   hmiStns[3].wip[6].pnCode[4] := 0;
   hmiStns[3].wip[6].pnCode[5] := 0;
   hmiStns[3].wip[6].pnCode[6] := 197000;
   hmiStns[3].wip[6].pnCode[7] := 179000;
   hmiStns[3].wip[7].wipCode := -1;
   hmiStns[3].wip[7].pnCode[0] := 0;
   hmiStns[3].wip[7].pnCode[1] := 243000;
   hmiStns[3].wip[7].pnCode[2] := 0;
   hmiStns[3].wip[7].pnCode[3] := 199000;
   hmiStns[3].wip[7].pnCode[4] := 0;
   hmiStns[3].wip[7].pnCode[5] := 0;
   hmiStns[3].wip[7].pnCode[6] := 198000;
   hmiStns[3].wip[7].pnCode[7] := 178000;
   hmiStns[3].wip[8].wipCode := -1;
   hmiStns[3].wip[8].pnCode[0] := 0;
   hmiStns[3].wip[8].pnCode[1] := 0;
   hmiStns[3].wip[8].pnCode[2] := 0;
   hmiStns[3].wip[8].pnCode[3] := 0;
   hmiStns[3].wip[8].pnCode[4] := 0;
   hmiStns[3].wip[8].pnCode[5] := 0;
   hmiStns[3].wip[8].pnCode[6] := 0;
   hmiStns[3].wip[8].pnCode[7] := 0;
   hmiStns[3].wip[9].wipCode := -1;
   hmiStns[3].wip[9].pnCode[0] := 0;
   hmiStns[3].wip[9].pnCode[1] := 0;
   hmiStns[3].wip[9].pnCode[2] := 0;
   hmiStns[3].wip[9].pnCode[3] := 0;
   hmiStns[3].wip[9].pnCode[4] := 0;
   hmiStns[3].wip[9].pnCode[5] := 0;
   hmiStns[3].wip[9].pnCode[6] := 0;
   hmiStns[3].wip[9].pnCode[7] := 0;
   hmiStns[3].wip[10].wipCode := -1;
   hmiStns[3].wip[10].pnCode[0] := 0;
   hmiStns[3].wip[10].pnCode[1] := 0;
   hmiStns[3].wip[10].pnCode[2] := 0;
   hmiStns[3].wip[10].pnCode[3] := 0;
   hmiStns[3].wip[10].pnCode[4] := 0;
   hmiStns[3].wip[10].pnCode[5] := 0;
   hmiStns[3].wip[10].pnCode[6] := 0;
   hmiStns[3].wip[10].pnCode[7] := 0;
   hmiStns[3].wip[11].wipCode := -1;
   hmiStns[3].wip[11].pnCode[0] := 0;
   hmiStns[3].wip[11].pnCode[1] := 0;
   hmiStns[3].wip[11].pnCode[2] := 0;
   hmiStns[3].wip[11].pnCode[3] := 0;
   hmiStns[3].wip[11].pnCode[4] := 0;
   hmiStns[3].wip[11].pnCode[5] := 0;
   hmiStns[3].wip[11].pnCode[6] := 0;
   hmiStns[3].wip[11].pnCode[7] := 0;
   hmiStns[3].wip[12].wipCode := -1;
   hmiStns[3].wip[12].pnCode[0] := 0;
   hmiStns[3].wip[12].pnCode[1] := 0;
   hmiStns[3].wip[12].pnCode[2] := 0;
   hmiStns[3].wip[12].pnCode[3] := 0;
   hmiStns[3].wip[12].pnCode[4] := 0;
   hmiStns[3].wip[12].pnCode[5] := 0;
   hmiStns[3].wip[12].pnCode[6] := 0;
   hmiStns[3].wip[12].pnCode[7] := 0;
   hmiStns[3].wip[13].wipCode := -1;
   hmiStns[3].wip[13].pnCode[0] := 0;
   hmiStns[3].wip[13].pnCode[1] := 0;
   hmiStns[3].wip[13].pnCode[2] := 0;
   hmiStns[3].wip[13].pnCode[3] := 0;
   hmiStns[3].wip[13].pnCode[4] := 0;
   hmiStns[3].wip[13].pnCode[5] := 0;
   hmiStns[3].wip[13].pnCode[6] := 0;
   hmiStns[3].wip[13].pnCode[7] := 0;
   hmiStns[3].wip[14].wipCode := -1;
   hmiStns[3].wip[14].pnCode[0] := 0;
   hmiStns[3].wip[14].pnCode[1] := 0;
   hmiStns[3].wip[14].pnCode[2] := 0;
   hmiStns[3].wip[14].pnCode[3] := 0;
   hmiStns[3].wip[14].pnCode[4] := 0;
   hmiStns[3].wip[14].pnCode[5] := 0;
   hmiStns[3].wip[14].pnCode[6] := 0;
   hmiStns[3].wip[14].pnCode[7] := 0;
   hmiStns[3].wip[15].wipCode := -1;
   hmiStns[3].wip[15].pnCode[0] := 0;
   hmiStns[3].wip[15].pnCode[1] := 0;
   hmiStns[3].wip[15].pnCode[2] := 0;
   hmiStns[3].wip[15].pnCode[3] := 0;
   hmiStns[3].wip[15].pnCode[4] := 0;
   hmiStns[3].wip[15].pnCode[5] := 0;
   hmiStns[3].wip[15].pnCode[6] := 0;
   hmiStns[3].wip[15].pnCode[7] := 0;
   hmiStns[3].wip[16].wipCode := -1;
   hmiStns[3].wip[16].pnCode[0] := 0;
   hmiStns[3].wip[16].pnCode[1] := 0;
   hmiStns[3].wip[16].pnCode[2] := 0;
   hmiStns[3].wip[16].pnCode[3] := 0;
   hmiStns[3].wip[16].pnCode[4] := 0;
   hmiStns[3].wip[16].pnCode[5] := 0;
   hmiStns[3].wip[16].pnCode[6] := 0;
   hmiStns[3].wip[16].pnCode[7] := 0;
   hmiStns[3].wip[17].wipCode := -1;
   hmiStns[3].wip[17].pnCode[0] := 0;
   hmiStns[3].wip[17].pnCode[1] := 0;
   hmiStns[3].wip[17].pnCode[2] := 0;
   hmiStns[3].wip[17].pnCode[3] := 0;
   hmiStns[3].wip[17].pnCode[4] := 0;
   hmiStns[3].wip[17].pnCode[5] := 0;
   hmiStns[3].wip[17].pnCode[6] := 0;
   hmiStns[3].wip[17].pnCode[7] := 0;
   hmiStns[3].wip[18].wipCode := -1;
   hmiStns[3].wip[18].pnCode[0] := 0;
   hmiStns[3].wip[18].pnCode[1] := 0;
   hmiStns[3].wip[18].pnCode[2] := 0;
   hmiStns[3].wip[18].pnCode[3] := 0;
   hmiStns[3].wip[18].pnCode[4] := 0;
   hmiStns[3].wip[18].pnCode[5] := 0;
   hmiStns[3].wip[18].pnCode[6] := 0;
   hmiStns[3].wip[18].pnCode[7] := 0;
   hmiStns[3].wip[19].wipCode := -1;
   hmiStns[3].wip[19].pnCode[0] := 0;
   hmiStns[3].wip[19].pnCode[1] := 0;
   hmiStns[3].wip[19].pnCode[2] := 0;
   hmiStns[3].wip[19].pnCode[3] := 0;
   hmiStns[3].wip[19].pnCode[4] := 0;
   hmiStns[3].wip[19].pnCode[5] := 0;
   hmiStns[3].wip[19].pnCode[6] := 0;
   hmiStns[3].wip[19].pnCode[7] := 0;
   hmiStns[3].wip[20].wipCode := -1;
   hmiStns[3].wip[20].pnCode[0] := 0;
   hmiStns[3].wip[20].pnCode[1] := 0;
   hmiStns[3].wip[20].pnCode[2] := 0;
   hmiStns[3].wip[20].pnCode[3] := 0;
   hmiStns[3].wip[20].pnCode[4] := 0;
   hmiStns[3].wip[20].pnCode[5] := 0;
   hmiStns[3].wip[20].pnCode[6] := 0;
   hmiStns[3].wip[20].pnCode[7] := 0;
   hmiStns[3].wip[21].wipCode := -1;
   hmiStns[3].wip[21].pnCode[0] := 0;
   hmiStns[3].wip[21].pnCode[1] := 0;
   hmiStns[3].wip[21].pnCode[2] := 0;
   hmiStns[3].wip[21].pnCode[3] := 0;
   hmiStns[3].wip[21].pnCode[4] := 0;
   hmiStns[3].wip[21].pnCode[5] := 0;
   hmiStns[3].wip[21].pnCode[6] := 0;
   hmiStns[3].wip[21].pnCode[7] := 0;
   hmiStns[3].wip[22].wipCode := -1;
   hmiStns[3].wip[22].pnCode[0] := 0;
   hmiStns[3].wip[22].pnCode[1] := 0;
   hmiStns[3].wip[22].pnCode[2] := 0;
   hmiStns[3].wip[22].pnCode[3] := 0;
   hmiStns[3].wip[22].pnCode[4] := 0;
   hmiStns[3].wip[22].pnCode[5] := 0;
   hmiStns[3].wip[22].pnCode[6] := 0;
   hmiStns[3].wip[22].pnCode[7] := 0;
   hmiStns[3].wip[23].wipCode := -1;
   hmiStns[3].wip[23].pnCode[0] := 0;
   hmiStns[3].wip[23].pnCode[1] := 0;
   hmiStns[3].wip[23].pnCode[2] := 0;
   hmiStns[3].wip[23].pnCode[3] := 0;
   hmiStns[3].wip[23].pnCode[4] := 0;
   hmiStns[3].wip[23].pnCode[5] := 0;
   hmiStns[3].wip[23].pnCode[6] := 0;
   hmiStns[3].wip[23].pnCode[7] := 0;
   hmiStns[3].wip[24].wipCode := -1;
   hmiStns[3].wip[24].pnCode[0] := 0;
   hmiStns[3].wip[24].pnCode[1] := 0;
   hmiStns[3].wip[24].pnCode[2] := 0;
   hmiStns[3].wip[24].pnCode[3] := 0;
   hmiStns[3].wip[24].pnCode[4] := 0;
   hmiStns[3].wip[24].pnCode[5] := 0;
   hmiStns[3].wip[24].pnCode[6] := 0;
   hmiStns[3].wip[24].pnCode[7] := 0;
   hmiStns[3].wip[25].wipCode := -1;
   hmiStns[3].wip[25].pnCode[0] := 0;
   hmiStns[3].wip[25].pnCode[1] := 0;
   hmiStns[3].wip[25].pnCode[2] := 0;
   hmiStns[3].wip[25].pnCode[3] := 0;
   hmiStns[3].wip[25].pnCode[4] := 0;
   hmiStns[3].wip[25].pnCode[5] := 0;
   hmiStns[3].wip[25].pnCode[6] := 0;
   hmiStns[3].wip[25].pnCode[7] := 0;
   hmiStns[3].wip[26].wipCode := -1;
   hmiStns[3].wip[26].pnCode[0] := 0;
   hmiStns[3].wip[26].pnCode[1] := 0;
   hmiStns[3].wip[26].pnCode[2] := 0;
   hmiStns[3].wip[26].pnCode[3] := 0;
   hmiStns[3].wip[26].pnCode[4] := 0;
   hmiStns[3].wip[26].pnCode[5] := 0;
   hmiStns[3].wip[26].pnCode[6] := 0;
   hmiStns[3].wip[26].pnCode[7] := 0;
   hmiStns[3].wip[27].wipCode := -1;
   hmiStns[3].wip[27].pnCode[0] := 0;
   hmiStns[3].wip[27].pnCode[1] := 0;
   hmiStns[3].wip[27].pnCode[2] := 0;
   hmiStns[3].wip[27].pnCode[3] := 0;
   hmiStns[3].wip[27].pnCode[4] := 0;
   hmiStns[3].wip[27].pnCode[5] := 0;
   hmiStns[3].wip[27].pnCode[6] := 0;
   hmiStns[3].wip[27].pnCode[7] := 0;
   hmiStns[3].wip[28].wipCode := -1;
   hmiStns[3].wip[28].pnCode[0] := 0;
   hmiStns[3].wip[28].pnCode[1] := 0;
   hmiStns[3].wip[28].pnCode[2] := 0;
   hmiStns[3].wip[28].pnCode[3] := 0;
   hmiStns[3].wip[28].pnCode[4] := 0;
   hmiStns[3].wip[28].pnCode[5] := 0;
   hmiStns[3].wip[28].pnCode[6] := 0;
   hmiStns[3].wip[28].pnCode[7] := 0;
   hmiStns[3].wip[29].wipCode := -1;
   hmiStns[3].wip[29].pnCode[0] := 0;
   hmiStns[3].wip[29].pnCode[1] := 0;
   hmiStns[3].wip[29].pnCode[2] := 0;
   hmiStns[3].wip[29].pnCode[3] := 0;
   hmiStns[3].wip[29].pnCode[4] := 0;
   hmiStns[3].wip[29].pnCode[5] := 0;
   hmiStns[3].wip[29].pnCode[6] := 0;
   hmiStns[3].wip[29].pnCode[7] := 0;
   hmiStns[3].wip[30].wipCode := -1;
   hmiStns[3].wip[30].pnCode[0] := 0;
   hmiStns[3].wip[30].pnCode[1] := 0;
   hmiStns[3].wip[30].pnCode[2] := 0;
   hmiStns[3].wip[30].pnCode[3] := 0;
   hmiStns[3].wip[30].pnCode[4] := 0;
   hmiStns[3].wip[30].pnCode[5] := 0;
   hmiStns[3].wip[30].pnCode[6] := 0;
   hmiStns[3].wip[30].pnCode[7] := 0;
   hmiStns[3].wip[31].wipCode := -1;
   hmiStns[3].wip[31].pnCode[0] := 0;
   hmiStns[3].wip[31].pnCode[1] := 0;
   hmiStns[3].wip[31].pnCode[2] := 0;
   hmiStns[3].wip[31].pnCode[3] := 0;
   hmiStns[3].wip[31].pnCode[4] := 0;
   hmiStns[3].wip[31].pnCode[5] := 0;
   hmiStns[3].wip[31].pnCode[6] := 0;
   hmiStns[3].wip[31].pnCode[7] := 0;
   hmiStns[3].wip[32].wipCode := -1;
   hmiStns[3].wip[32].pnCode[0] := 0;
   hmiStns[3].wip[32].pnCode[1] := 0;
   hmiStns[3].wip[32].pnCode[2] := 0;
   hmiStns[3].wip[32].pnCode[3] := 0;
   hmiStns[3].wip[32].pnCode[4] := 0;
   hmiStns[3].wip[32].pnCode[5] := 0;
   hmiStns[3].wip[32].pnCode[6] := 0;
   hmiStns[3].wip[32].pnCode[7] := 0;
   hmiStns[3].wip[33].wipCode := -1;
   hmiStns[3].wip[33].pnCode[0] := 0;
   hmiStns[3].wip[33].pnCode[1] := 0;
   hmiStns[3].wip[33].pnCode[2] := 0;
   hmiStns[3].wip[33].pnCode[3] := 0;
   hmiStns[3].wip[33].pnCode[4] := 0;
   hmiStns[3].wip[33].pnCode[5] := 0;
   hmiStns[3].wip[33].pnCode[6] := 0;
   hmiStns[3].wip[33].pnCode[7] := 0;
   hmiStns[3].wip[34].wipCode := -1;
   hmiStns[3].wip[34].pnCode[0] := 0;
   hmiStns[3].wip[34].pnCode[1] := 0;
   hmiStns[3].wip[34].pnCode[2] := 0;
   hmiStns[3].wip[34].pnCode[3] := 0;
   hmiStns[3].wip[34].pnCode[4] := 0;
   hmiStns[3].wip[34].pnCode[5] := 0;
   hmiStns[3].wip[34].pnCode[6] := 0;
   hmiStns[3].wip[34].pnCode[7] := 0;
   hmiStns[3].wip[35].wipCode := -1;
   hmiStns[3].wip[35].pnCode[0] := 0;
   hmiStns[3].wip[35].pnCode[1] := 0;
   hmiStns[3].wip[35].pnCode[2] := 0;
   hmiStns[3].wip[35].pnCode[3] := 0;
   hmiStns[3].wip[35].pnCode[4] := 0;
   hmiStns[3].wip[35].pnCode[5] := 0;
   hmiStns[3].wip[35].pnCode[6] := 0;
   hmiStns[3].wip[35].pnCode[7] := 0;
   hmiStns[3].wip[36].wipCode := -1;
   hmiStns[3].wip[36].pnCode[0] := 0;
   hmiStns[3].wip[36].pnCode[1] := 0;
   hmiStns[3].wip[36].pnCode[2] := 0;
   hmiStns[3].wip[36].pnCode[3] := 0;
   hmiStns[3].wip[36].pnCode[4] := 0;
   hmiStns[3].wip[36].pnCode[5] := 0;
   hmiStns[3].wip[36].pnCode[6] := 0;
   hmiStns[3].wip[36].pnCode[7] := 0;
   hmiStns[3].wip[37].wipCode := -1;
   hmiStns[3].wip[37].pnCode[0] := 0;
   hmiStns[3].wip[37].pnCode[1] := 0;
   hmiStns[3].wip[37].pnCode[2] := 0;
   hmiStns[3].wip[37].pnCode[3] := 0;
   hmiStns[3].wip[37].pnCode[4] := 0;
   hmiStns[3].wip[37].pnCode[5] := 0;
   hmiStns[3].wip[37].pnCode[6] := 0;
   hmiStns[3].wip[37].pnCode[7] := 0;
   hmiStns[3].wip[38].wipCode := -1;
   hmiStns[3].wip[38].pnCode[0] := 0;
   hmiStns[3].wip[38].pnCode[1] := 0;
   hmiStns[3].wip[38].pnCode[2] := 0;
   hmiStns[3].wip[38].pnCode[3] := 0;
   hmiStns[3].wip[38].pnCode[4] := 0;
   hmiStns[3].wip[38].pnCode[5] := 0;
   hmiStns[3].wip[38].pnCode[6] := 0;
   hmiStns[3].wip[38].pnCode[7] := 0;
   hmiStns[3].wip[39].wipCode := -1;
   hmiStns[3].wip[39].pnCode[0] := 0;
   hmiStns[3].wip[39].pnCode[1] := 0;
   hmiStns[3].wip[39].pnCode[2] := 0;
   hmiStns[3].wip[39].pnCode[3] := 0;
   hmiStns[3].wip[39].pnCode[4] := 0;
   hmiStns[3].wip[39].pnCode[5] := 0;
   hmiStns[3].wip[39].pnCode[6] := 0;
   hmiStns[3].wip[39].pnCode[7] := 0;
   hmiStns[3].wip[40].wipCode := -1;
   hmiStns[3].wip[40].pnCode[0] := 0;
   hmiStns[3].wip[40].pnCode[1] := 0;
   hmiStns[3].wip[40].pnCode[2] := 0;
   hmiStns[3].wip[40].pnCode[3] := 0;
   hmiStns[3].wip[40].pnCode[4] := 0;
   hmiStns[3].wip[40].pnCode[5] := 0;
   hmiStns[3].wip[40].pnCode[6] := 0;
   hmiStns[3].wip[40].pnCode[7] := 0;
   hmiStns[3].wip[41].wipCode := -1;
   hmiStns[3].wip[41].pnCode[0] := 0;
   hmiStns[3].wip[41].pnCode[1] := 0;
   hmiStns[3].wip[41].pnCode[2] := 0;
   hmiStns[3].wip[41].pnCode[3] := 0;
   hmiStns[3].wip[41].pnCode[4] := 0;
   hmiStns[3].wip[41].pnCode[5] := 0;
   hmiStns[3].wip[41].pnCode[6] := 0;
   hmiStns[3].wip[41].pnCode[7] := 0;
   hmiStns[3].wip[42].wipCode := -1;
   hmiStns[3].wip[42].pnCode[0] := 0;
   hmiStns[3].wip[42].pnCode[1] := 0;
   hmiStns[3].wip[42].pnCode[2] := 0;
   hmiStns[3].wip[42].pnCode[3] := 0;
   hmiStns[3].wip[42].pnCode[4] := 0;
   hmiStns[3].wip[42].pnCode[5] := 0;
   hmiStns[3].wip[42].pnCode[6] := 0;
   hmiStns[3].wip[42].pnCode[7] := 0;
   hmiStns[3].wip[43].wipCode := -1;
   hmiStns[3].wip[43].pnCode[0] := 0;
   hmiStns[3].wip[43].pnCode[1] := 0;
   hmiStns[3].wip[43].pnCode[2] := 0;
   hmiStns[3].wip[43].pnCode[3] := 0;
   hmiStns[3].wip[43].pnCode[4] := 0;
   hmiStns[3].wip[43].pnCode[5] := 0;
   hmiStns[3].wip[43].pnCode[6] := 0;
   hmiStns[3].wip[43].pnCode[7] := 0;
   hmiStns[3].wip[44].wipCode := -1;
   hmiStns[3].wip[44].pnCode[0] := 0;
   hmiStns[3].wip[44].pnCode[1] := 0;
   hmiStns[3].wip[44].pnCode[2] := 0;
   hmiStns[3].wip[44].pnCode[3] := 0;
   hmiStns[3].wip[44].pnCode[4] := 0;
   hmiStns[3].wip[44].pnCode[5] := 0;
   hmiStns[3].wip[44].pnCode[6] := 0;
   hmiStns[3].wip[44].pnCode[7] := 0;
   hmiStns[3].wip[45].wipCode := -1;
   hmiStns[3].wip[45].pnCode[0] := 0;
   hmiStns[3].wip[45].pnCode[1] := 0;
   hmiStns[3].wip[45].pnCode[2] := 0;
   hmiStns[3].wip[45].pnCode[3] := 0;
   hmiStns[3].wip[45].pnCode[4] := 0;
   hmiStns[3].wip[45].pnCode[5] := 0;
   hmiStns[3].wip[45].pnCode[6] := 0;
   hmiStns[3].wip[45].pnCode[7] := 0;
   hmiStns[3].wip[46].wipCode := -1;
   hmiStns[3].wip[46].pnCode[0] := 0;
   hmiStns[3].wip[46].pnCode[1] := 0;
   hmiStns[3].wip[46].pnCode[2] := 0;
   hmiStns[3].wip[46].pnCode[3] := 0;
   hmiStns[3].wip[46].pnCode[4] := 0;
   hmiStns[3].wip[46].pnCode[5] := 0;
   hmiStns[3].wip[46].pnCode[6] := 0;
   hmiStns[3].wip[46].pnCode[7] := 0;
   hmiStns[3].wip[47].wipCode := -1;
   hmiStns[3].wip[47].pnCode[0] := 0;
   hmiStns[3].wip[47].pnCode[1] := 0;
   hmiStns[3].wip[47].pnCode[2] := 0;
   hmiStns[3].wip[47].pnCode[3] := 0;
   hmiStns[3].wip[47].pnCode[4] := 0;
   hmiStns[3].wip[47].pnCode[5] := 0;
   hmiStns[3].wip[47].pnCode[6] := 0;
   hmiStns[3].wip[47].pnCode[7] := 0;
   hmiStns[3].wip[48].wipCode := -1;
   hmiStns[3].wip[48].pnCode[0] := 0;
   hmiStns[3].wip[48].pnCode[1] := 0;
   hmiStns[3].wip[48].pnCode[2] := 0;
   hmiStns[3].wip[48].pnCode[3] := 0;
   hmiStns[3].wip[48].pnCode[4] := 0;
   hmiStns[3].wip[48].pnCode[5] := 0;
   hmiStns[3].wip[48].pnCode[6] := 0;
   hmiStns[3].wip[48].pnCode[7] := 0;
   hmiStns[3].wip[49].wipCode := -1;
   hmiStns[3].wip[49].pnCode[0] := 0;
   hmiStns[3].wip[49].pnCode[1] := 0;
   hmiStns[3].wip[49].pnCode[2] := 0;
   hmiStns[3].wip[49].pnCode[3] := 0;
   hmiStns[3].wip[49].pnCode[4] := 0;
   hmiStns[3].wip[49].pnCode[5] := 0;
   hmiStns[3].wip[49].pnCode[6] := 0;
   hmiStns[3].wip[49].pnCode[7] := 0;
   hmiStns[4].wip[0].wipCode := 1032;
   hmiStns[4].wip[0].pnCode[0] := 0;
   hmiStns[4].wip[0].pnCode[1] := 243000;
   hmiStns[4].wip[0].pnCode[2] := 0;
   hmiStns[4].wip[0].pnCode[3] := 3000;
   hmiStns[4].wip[0].pnCode[4] := 0;
   hmiStns[4].wip[0].pnCode[5] := 0;
   hmiStns[4].wip[0].pnCode[6] := 1000;
   hmiStns[4].wip[0].pnCode[7] := 2000;
   hmiStns[4].wip[1].wipCode := 2059;
   hmiStns[4].wip[1].pnCode[0] := 0;
   hmiStns[4].wip[1].pnCode[1] := 243000;
   hmiStns[4].wip[1].pnCode[2] := 5000;
   hmiStns[4].wip[1].pnCode[3] := 9000;
   hmiStns[4].wip[1].pnCode[4] := 0;
   hmiStns[4].wip[1].pnCode[5] := 6000;
   hmiStns[4].wip[1].pnCode[6] := 4000;
   hmiStns[4].wip[1].pnCode[7] := 10000;
   hmiStns[4].wip[2].wipCode := 3059;
   hmiStns[4].wip[2].pnCode[0] := 0;
   hmiStns[4].wip[2].pnCode[1] := 243000;
   hmiStns[4].wip[2].pnCode[2] := 7000;
   hmiStns[4].wip[2].pnCode[3] := 9000;
   hmiStns[4].wip[2].pnCode[4] := 0;
   hmiStns[4].wip[2].pnCode[5] := 8000;
   hmiStns[4].wip[2].pnCode[6] := 4000;
   hmiStns[4].wip[2].pnCode[7] := 10000;
   hmiStns[4].wip[3].wipCode := -1;
   hmiStns[4].wip[3].pnCode[0] := 0;
   hmiStns[4].wip[3].pnCode[1] := 0;
   hmiStns[4].wip[3].pnCode[2] := 0;
   hmiStns[4].wip[3].pnCode[3] := 0;
   hmiStns[4].wip[3].pnCode[4] := 0;
   hmiStns[4].wip[3].pnCode[5] := 0;
   hmiStns[4].wip[3].pnCode[6] := 0;
   hmiStns[4].wip[3].pnCode[7] := 0;
   hmiStns[4].wip[4].wipCode := -1;
   hmiStns[4].wip[4].pnCode[0] := 0;
   hmiStns[4].wip[4].pnCode[1] := 0;
   hmiStns[4].wip[4].pnCode[2] := 0;
   hmiStns[4].wip[4].pnCode[3] := 0;
   hmiStns[4].wip[4].pnCode[4] := 0;
   hmiStns[4].wip[4].pnCode[5] := 0;
   hmiStns[4].wip[4].pnCode[6] := 0;
   hmiStns[4].wip[4].pnCode[7] := 0;
   hmiStns[4].wip[5].wipCode := -1;
   hmiStns[4].wip[5].pnCode[0] := 0;
   hmiStns[4].wip[5].pnCode[1] := 0;
   hmiStns[4].wip[5].pnCode[2] := 0;
   hmiStns[4].wip[5].pnCode[3] := 0;
   hmiStns[4].wip[5].pnCode[4] := 0;
   hmiStns[4].wip[5].pnCode[5] := 0;
   hmiStns[4].wip[5].pnCode[6] := 0;
   hmiStns[4].wip[5].pnCode[7] := 0;
   hmiStns[4].wip[6].wipCode := -1;
   hmiStns[4].wip[6].pnCode[0] := 0;
   hmiStns[4].wip[6].pnCode[1] := 0;
   hmiStns[4].wip[6].pnCode[2] := 0;
   hmiStns[4].wip[6].pnCode[3] := 0;
   hmiStns[4].wip[6].pnCode[4] := 0;
   hmiStns[4].wip[6].pnCode[5] := 0;
   hmiStns[4].wip[6].pnCode[6] := 0;
   hmiStns[4].wip[6].pnCode[7] := 0;
   hmiStns[4].wip[7].wipCode := -1;
   hmiStns[4].wip[7].pnCode[0] := 0;
   hmiStns[4].wip[7].pnCode[1] := 0;
   hmiStns[4].wip[7].pnCode[2] := 0;
   hmiStns[4].wip[7].pnCode[3] := 0;
   hmiStns[4].wip[7].pnCode[4] := 0;
   hmiStns[4].wip[7].pnCode[5] := 0;
   hmiStns[4].wip[7].pnCode[6] := 0;
   hmiStns[4].wip[7].pnCode[7] := 0;
   hmiStns[4].wip[8].wipCode := -1;
   hmiStns[4].wip[8].pnCode[0] := 0;
   hmiStns[4].wip[8].pnCode[1] := 0;
   hmiStns[4].wip[8].pnCode[2] := 0;
   hmiStns[4].wip[8].pnCode[3] := 0;
   hmiStns[4].wip[8].pnCode[4] := 0;
   hmiStns[4].wip[8].pnCode[5] := 0;
   hmiStns[4].wip[8].pnCode[6] := 0;
   hmiStns[4].wip[8].pnCode[7] := 0;
   hmiStns[4].wip[9].wipCode := -1;
   hmiStns[4].wip[9].pnCode[0] := 0;
   hmiStns[4].wip[9].pnCode[1] := 0;
   hmiStns[4].wip[9].pnCode[2] := 0;
   hmiStns[4].wip[9].pnCode[3] := 0;
   hmiStns[4].wip[9].pnCode[4] := 0;
   hmiStns[4].wip[9].pnCode[5] := 0;
   hmiStns[4].wip[9].pnCode[6] := 0;
   hmiStns[4].wip[9].pnCode[7] := 0;
   hmiStns[4].wip[10].wipCode := -1;
   hmiStns[4].wip[10].pnCode[0] := 0;
   hmiStns[4].wip[10].pnCode[1] := 0;
   hmiStns[4].wip[10].pnCode[2] := 0;
   hmiStns[4].wip[10].pnCode[3] := 0;
   hmiStns[4].wip[10].pnCode[4] := 0;
   hmiStns[4].wip[10].pnCode[5] := 0;
   hmiStns[4].wip[10].pnCode[6] := 0;
   hmiStns[4].wip[10].pnCode[7] := 0;
   hmiStns[4].wip[11].wipCode := -1;
   hmiStns[4].wip[11].pnCode[0] := 0;
   hmiStns[4].wip[11].pnCode[1] := 0;
   hmiStns[4].wip[11].pnCode[2] := 0;
   hmiStns[4].wip[11].pnCode[3] := 0;
   hmiStns[4].wip[11].pnCode[4] := 0;
   hmiStns[4].wip[11].pnCode[5] := 0;
   hmiStns[4].wip[11].pnCode[6] := 0;
   hmiStns[4].wip[11].pnCode[7] := 0;
   hmiStns[4].wip[12].wipCode := -1;
   hmiStns[4].wip[12].pnCode[0] := 0;
   hmiStns[4].wip[12].pnCode[1] := 0;
   hmiStns[4].wip[12].pnCode[2] := 0;
   hmiStns[4].wip[12].pnCode[3] := 0;
   hmiStns[4].wip[12].pnCode[4] := 0;
   hmiStns[4].wip[12].pnCode[5] := 0;
   hmiStns[4].wip[12].pnCode[6] := 0;
   hmiStns[4].wip[12].pnCode[7] := 0;
   hmiStns[4].wip[13].wipCode := -1;
   hmiStns[4].wip[13].pnCode[0] := 0;
   hmiStns[4].wip[13].pnCode[1] := 0;
   hmiStns[4].wip[13].pnCode[2] := 0;
   hmiStns[4].wip[13].pnCode[3] := 0;
   hmiStns[4].wip[13].pnCode[4] := 0;
   hmiStns[4].wip[13].pnCode[5] := 0;
   hmiStns[4].wip[13].pnCode[6] := 0;
   hmiStns[4].wip[13].pnCode[7] := 0;
   hmiStns[4].wip[14].wipCode := -1;
   hmiStns[4].wip[14].pnCode[0] := 0;
   hmiStns[4].wip[14].pnCode[1] := 0;
   hmiStns[4].wip[14].pnCode[2] := 0;
   hmiStns[4].wip[14].pnCode[3] := 0;
   hmiStns[4].wip[14].pnCode[4] := 0;
   hmiStns[4].wip[14].pnCode[5] := 0;
   hmiStns[4].wip[14].pnCode[6] := 0;
   hmiStns[4].wip[14].pnCode[7] := 0;
   hmiStns[4].wip[15].wipCode := -1;
   hmiStns[4].wip[15].pnCode[0] := 0;
   hmiStns[4].wip[15].pnCode[1] := 0;
   hmiStns[4].wip[15].pnCode[2] := 0;
   hmiStns[4].wip[15].pnCode[3] := 0;
   hmiStns[4].wip[15].pnCode[4] := 0;
   hmiStns[4].wip[15].pnCode[5] := 0;
   hmiStns[4].wip[15].pnCode[6] := 0;
   hmiStns[4].wip[15].pnCode[7] := 0;
   hmiStns[4].wip[16].wipCode := -1;
   hmiStns[4].wip[16].pnCode[0] := 0;
   hmiStns[4].wip[16].pnCode[1] := 0;
   hmiStns[4].wip[16].pnCode[2] := 0;
   hmiStns[4].wip[16].pnCode[3] := 0;
   hmiStns[4].wip[16].pnCode[4] := 0;
   hmiStns[4].wip[16].pnCode[5] := 0;
   hmiStns[4].wip[16].pnCode[6] := 0;
   hmiStns[4].wip[16].pnCode[7] := 0;
   hmiStns[4].wip[17].wipCode := -1;
   hmiStns[4].wip[17].pnCode[0] := 0;
   hmiStns[4].wip[17].pnCode[1] := 0;
   hmiStns[4].wip[17].pnCode[2] := 0;
   hmiStns[4].wip[17].pnCode[3] := 0;
   hmiStns[4].wip[17].pnCode[4] := 0;
   hmiStns[4].wip[17].pnCode[5] := 0;
   hmiStns[4].wip[17].pnCode[6] := 0;
   hmiStns[4].wip[17].pnCode[7] := 0;
   hmiStns[4].wip[18].wipCode := -1;
   hmiStns[4].wip[18].pnCode[0] := 0;
   hmiStns[4].wip[18].pnCode[1] := 0;
   hmiStns[4].wip[18].pnCode[2] := 0;
   hmiStns[4].wip[18].pnCode[3] := 0;
   hmiStns[4].wip[18].pnCode[4] := 0;
   hmiStns[4].wip[18].pnCode[5] := 0;
   hmiStns[4].wip[18].pnCode[6] := 0;
   hmiStns[4].wip[18].pnCode[7] := 0;
   hmiStns[4].wip[19].wipCode := -1;
   hmiStns[4].wip[19].pnCode[0] := 0;
   hmiStns[4].wip[19].pnCode[1] := 0;
   hmiStns[4].wip[19].pnCode[2] := 0;
   hmiStns[4].wip[19].pnCode[3] := 0;
   hmiStns[4].wip[19].pnCode[4] := 0;
   hmiStns[4].wip[19].pnCode[5] := 0;
   hmiStns[4].wip[19].pnCode[6] := 0;
   hmiStns[4].wip[19].pnCode[7] := 0;
   hmiStns[4].wip[20].wipCode := -1;
   hmiStns[4].wip[20].pnCode[0] := 0;
   hmiStns[4].wip[20].pnCode[1] := 0;
   hmiStns[4].wip[20].pnCode[2] := 0;
   hmiStns[4].wip[20].pnCode[3] := 0;
   hmiStns[4].wip[20].pnCode[4] := 0;
   hmiStns[4].wip[20].pnCode[5] := 0;
   hmiStns[4].wip[20].pnCode[6] := 0;
   hmiStns[4].wip[20].pnCode[7] := 0;
   hmiStns[4].wip[21].wipCode := -1;
   hmiStns[4].wip[21].pnCode[0] := 0;
   hmiStns[4].wip[21].pnCode[1] := 0;
   hmiStns[4].wip[21].pnCode[2] := 0;
   hmiStns[4].wip[21].pnCode[3] := 0;
   hmiStns[4].wip[21].pnCode[4] := 0;
   hmiStns[4].wip[21].pnCode[5] := 0;
   hmiStns[4].wip[21].pnCode[6] := 0;
   hmiStns[4].wip[21].pnCode[7] := 0;
   hmiStns[4].wip[22].wipCode := -1;
   hmiStns[4].wip[22].pnCode[0] := 0;
   hmiStns[4].wip[22].pnCode[1] := 0;
   hmiStns[4].wip[22].pnCode[2] := 0;
   hmiStns[4].wip[22].pnCode[3] := 0;
   hmiStns[4].wip[22].pnCode[4] := 0;
   hmiStns[4].wip[22].pnCode[5] := 0;
   hmiStns[4].wip[22].pnCode[6] := 0;
   hmiStns[4].wip[22].pnCode[7] := 0;
   hmiStns[4].wip[23].wipCode := -1;
   hmiStns[4].wip[23].pnCode[0] := 0;
   hmiStns[4].wip[23].pnCode[1] := 0;
   hmiStns[4].wip[23].pnCode[2] := 0;
   hmiStns[4].wip[23].pnCode[3] := 0;
   hmiStns[4].wip[23].pnCode[4] := 0;
   hmiStns[4].wip[23].pnCode[5] := 0;
   hmiStns[4].wip[23].pnCode[6] := 0;
   hmiStns[4].wip[23].pnCode[7] := 0;
   hmiStns[4].wip[24].wipCode := -1;
   hmiStns[4].wip[24].pnCode[0] := 0;
   hmiStns[4].wip[24].pnCode[1] := 0;
   hmiStns[4].wip[24].pnCode[2] := 0;
   hmiStns[4].wip[24].pnCode[3] := 0;
   hmiStns[4].wip[24].pnCode[4] := 0;
   hmiStns[4].wip[24].pnCode[5] := 0;
   hmiStns[4].wip[24].pnCode[6] := 0;
   hmiStns[4].wip[24].pnCode[7] := 0;
   hmiStns[4].wip[25].wipCode := -1;
   hmiStns[4].wip[25].pnCode[0] := 0;
   hmiStns[4].wip[25].pnCode[1] := 0;
   hmiStns[4].wip[25].pnCode[2] := 0;
   hmiStns[4].wip[25].pnCode[3] := 0;
   hmiStns[4].wip[25].pnCode[4] := 0;
   hmiStns[4].wip[25].pnCode[5] := 0;
   hmiStns[4].wip[25].pnCode[6] := 0;
   hmiStns[4].wip[25].pnCode[7] := 0;
   hmiStns[4].wip[26].wipCode := -1;
   hmiStns[4].wip[26].pnCode[0] := 0;
   hmiStns[4].wip[26].pnCode[1] := 0;
   hmiStns[4].wip[26].pnCode[2] := 0;
   hmiStns[4].wip[26].pnCode[3] := 0;
   hmiStns[4].wip[26].pnCode[4] := 0;
   hmiStns[4].wip[26].pnCode[5] := 0;
   hmiStns[4].wip[26].pnCode[6] := 0;
   hmiStns[4].wip[26].pnCode[7] := 0;
   hmiStns[4].wip[27].wipCode := -1;
   hmiStns[4].wip[27].pnCode[0] := 0;
   hmiStns[4].wip[27].pnCode[1] := 0;
   hmiStns[4].wip[27].pnCode[2] := 0;
   hmiStns[4].wip[27].pnCode[3] := 0;
   hmiStns[4].wip[27].pnCode[4] := 0;
   hmiStns[4].wip[27].pnCode[5] := 0;
   hmiStns[4].wip[27].pnCode[6] := 0;
   hmiStns[4].wip[27].pnCode[7] := 0;
   hmiStns[4].wip[28].wipCode := -1;
   hmiStns[4].wip[28].pnCode[0] := 0;
   hmiStns[4].wip[28].pnCode[1] := 0;
   hmiStns[4].wip[28].pnCode[2] := 0;
   hmiStns[4].wip[28].pnCode[3] := 0;
   hmiStns[4].wip[28].pnCode[4] := 0;
   hmiStns[4].wip[28].pnCode[5] := 0;
   hmiStns[4].wip[28].pnCode[6] := 0;
   hmiStns[4].wip[28].pnCode[7] := 0;
   hmiStns[4].wip[29].wipCode := -1;
   hmiStns[4].wip[29].pnCode[0] := 0;
   hmiStns[4].wip[29].pnCode[1] := 0;
   hmiStns[4].wip[29].pnCode[2] := 0;
   hmiStns[4].wip[29].pnCode[3] := 0;
   hmiStns[4].wip[29].pnCode[4] := 0;
   hmiStns[4].wip[29].pnCode[5] := 0;
   hmiStns[4].wip[29].pnCode[6] := 0;
   hmiStns[4].wip[29].pnCode[7] := 0;
   hmiStns[4].wip[30].wipCode := -1;
   hmiStns[4].wip[30].pnCode[0] := 0;
   hmiStns[4].wip[30].pnCode[1] := 0;
   hmiStns[4].wip[30].pnCode[2] := 0;
   hmiStns[4].wip[30].pnCode[3] := 0;
   hmiStns[4].wip[30].pnCode[4] := 0;
   hmiStns[4].wip[30].pnCode[5] := 0;
   hmiStns[4].wip[30].pnCode[6] := 0;
   hmiStns[4].wip[30].pnCode[7] := 0;
   hmiStns[4].wip[31].wipCode := -1;
   hmiStns[4].wip[31].pnCode[0] := 0;
   hmiStns[4].wip[31].pnCode[1] := 0;
   hmiStns[4].wip[31].pnCode[2] := 0;
   hmiStns[4].wip[31].pnCode[3] := 0;
   hmiStns[4].wip[31].pnCode[4] := 0;
   hmiStns[4].wip[31].pnCode[5] := 0;
   hmiStns[4].wip[31].pnCode[6] := 0;
   hmiStns[4].wip[31].pnCode[7] := 0;
   hmiStns[4].wip[32].wipCode := -1;
   hmiStns[4].wip[32].pnCode[0] := 0;
   hmiStns[4].wip[32].pnCode[1] := 0;
   hmiStns[4].wip[32].pnCode[2] := 0;
   hmiStns[4].wip[32].pnCode[3] := 0;
   hmiStns[4].wip[32].pnCode[4] := 0;
   hmiStns[4].wip[32].pnCode[5] := 0;
   hmiStns[4].wip[32].pnCode[6] := 0;
   hmiStns[4].wip[32].pnCode[7] := 0;
   hmiStns[4].wip[33].wipCode := -1;
   hmiStns[4].wip[33].pnCode[0] := 0;
   hmiStns[4].wip[33].pnCode[1] := 0;
   hmiStns[4].wip[33].pnCode[2] := 0;
   hmiStns[4].wip[33].pnCode[3] := 0;
   hmiStns[4].wip[33].pnCode[4] := 0;
   hmiStns[4].wip[33].pnCode[5] := 0;
   hmiStns[4].wip[33].pnCode[6] := 0;
   hmiStns[4].wip[33].pnCode[7] := 0;
   hmiStns[4].wip[34].wipCode := -1;
   hmiStns[4].wip[34].pnCode[0] := 0;
   hmiStns[4].wip[34].pnCode[1] := 0;
   hmiStns[4].wip[34].pnCode[2] := 0;
   hmiStns[4].wip[34].pnCode[3] := 0;
   hmiStns[4].wip[34].pnCode[4] := 0;
   hmiStns[4].wip[34].pnCode[5] := 0;
   hmiStns[4].wip[34].pnCode[6] := 0;
   hmiStns[4].wip[34].pnCode[7] := 0;
   hmiStns[4].wip[35].wipCode := -1;
   hmiStns[4].wip[35].pnCode[0] := 0;
   hmiStns[4].wip[35].pnCode[1] := 0;
   hmiStns[4].wip[35].pnCode[2] := 0;
   hmiStns[4].wip[35].pnCode[3] := 0;
   hmiStns[4].wip[35].pnCode[4] := 0;
   hmiStns[4].wip[35].pnCode[5] := 0;
   hmiStns[4].wip[35].pnCode[6] := 0;
   hmiStns[4].wip[35].pnCode[7] := 0;
   hmiStns[4].wip[36].wipCode := -1;
   hmiStns[4].wip[36].pnCode[0] := 0;
   hmiStns[4].wip[36].pnCode[1] := 0;
   hmiStns[4].wip[36].pnCode[2] := 0;
   hmiStns[4].wip[36].pnCode[3] := 0;
   hmiStns[4].wip[36].pnCode[4] := 0;
   hmiStns[4].wip[36].pnCode[5] := 0;
   hmiStns[4].wip[36].pnCode[6] := 0;
   hmiStns[4].wip[36].pnCode[7] := 0;
   hmiStns[4].wip[37].wipCode := -1;
   hmiStns[4].wip[37].pnCode[0] := 0;
   hmiStns[4].wip[37].pnCode[1] := 0;
   hmiStns[4].wip[37].pnCode[2] := 0;
   hmiStns[4].wip[37].pnCode[3] := 0;
   hmiStns[4].wip[37].pnCode[4] := 0;
   hmiStns[4].wip[37].pnCode[5] := 0;
   hmiStns[4].wip[37].pnCode[6] := 0;
   hmiStns[4].wip[37].pnCode[7] := 0;
   hmiStns[4].wip[38].wipCode := -1;
   hmiStns[4].wip[38].pnCode[0] := 0;
   hmiStns[4].wip[38].pnCode[1] := 0;
   hmiStns[4].wip[38].pnCode[2] := 0;
   hmiStns[4].wip[38].pnCode[3] := 0;
   hmiStns[4].wip[38].pnCode[4] := 0;
   hmiStns[4].wip[38].pnCode[5] := 0;
   hmiStns[4].wip[38].pnCode[6] := 0;
   hmiStns[4].wip[38].pnCode[7] := 0;
   hmiStns[4].wip[39].wipCode := -1;
   hmiStns[4].wip[39].pnCode[0] := 0;
   hmiStns[4].wip[39].pnCode[1] := 0;
   hmiStns[4].wip[39].pnCode[2] := 0;
   hmiStns[4].wip[39].pnCode[3] := 0;
   hmiStns[4].wip[39].pnCode[4] := 0;
   hmiStns[4].wip[39].pnCode[5] := 0;
   hmiStns[4].wip[39].pnCode[6] := 0;
   hmiStns[4].wip[39].pnCode[7] := 0;
   hmiStns[4].wip[40].wipCode := -1;
   hmiStns[4].wip[40].pnCode[0] := 0;
   hmiStns[4].wip[40].pnCode[1] := 0;
   hmiStns[4].wip[40].pnCode[2] := 0;
   hmiStns[4].wip[40].pnCode[3] := 0;
   hmiStns[4].wip[40].pnCode[4] := 0;
   hmiStns[4].wip[40].pnCode[5] := 0;
   hmiStns[4].wip[40].pnCode[6] := 0;
   hmiStns[4].wip[40].pnCode[7] := 0;
   hmiStns[4].wip[41].wipCode := -1;
   hmiStns[4].wip[41].pnCode[0] := 0;
   hmiStns[4].wip[41].pnCode[1] := 0;
   hmiStns[4].wip[41].pnCode[2] := 0;
   hmiStns[4].wip[41].pnCode[3] := 0;
   hmiStns[4].wip[41].pnCode[4] := 0;
   hmiStns[4].wip[41].pnCode[5] := 0;
   hmiStns[4].wip[41].pnCode[6] := 0;
   hmiStns[4].wip[41].pnCode[7] := 0;
   hmiStns[4].wip[42].wipCode := -1;
   hmiStns[4].wip[42].pnCode[0] := 0;
   hmiStns[4].wip[42].pnCode[1] := 0;
   hmiStns[4].wip[42].pnCode[2] := 0;
   hmiStns[4].wip[42].pnCode[3] := 0;
   hmiStns[4].wip[42].pnCode[4] := 0;
   hmiStns[4].wip[42].pnCode[5] := 0;
   hmiStns[4].wip[42].pnCode[6] := 0;
   hmiStns[4].wip[42].pnCode[7] := 0;
   hmiStns[4].wip[43].wipCode := -1;
   hmiStns[4].wip[43].pnCode[0] := 0;
   hmiStns[4].wip[43].pnCode[1] := 0;
   hmiStns[4].wip[43].pnCode[2] := 0;
   hmiStns[4].wip[43].pnCode[3] := 0;
   hmiStns[4].wip[43].pnCode[4] := 0;
   hmiStns[4].wip[43].pnCode[5] := 0;
   hmiStns[4].wip[43].pnCode[6] := 0;
   hmiStns[4].wip[43].pnCode[7] := 0;
   hmiStns[4].wip[44].wipCode := -1;
   hmiStns[4].wip[44].pnCode[0] := 0;
   hmiStns[4].wip[44].pnCode[1] := 0;
   hmiStns[4].wip[44].pnCode[2] := 0;
   hmiStns[4].wip[44].pnCode[3] := 0;
   hmiStns[4].wip[44].pnCode[4] := 0;
   hmiStns[4].wip[44].pnCode[5] := 0;
   hmiStns[4].wip[44].pnCode[6] := 0;
   hmiStns[4].wip[44].pnCode[7] := 0;
   hmiStns[4].wip[45].wipCode := -1;
   hmiStns[4].wip[45].pnCode[0] := 0;
   hmiStns[4].wip[45].pnCode[1] := 0;
   hmiStns[4].wip[45].pnCode[2] := 0;
   hmiStns[4].wip[45].pnCode[3] := 0;
   hmiStns[4].wip[45].pnCode[4] := 0;
   hmiStns[4].wip[45].pnCode[5] := 0;
   hmiStns[4].wip[45].pnCode[6] := 0;
   hmiStns[4].wip[45].pnCode[7] := 0;
   hmiStns[4].wip[46].wipCode := -1;
   hmiStns[4].wip[46].pnCode[0] := 0;
   hmiStns[4].wip[46].pnCode[1] := 0;
   hmiStns[4].wip[46].pnCode[2] := 0;
   hmiStns[4].wip[46].pnCode[3] := 0;
   hmiStns[4].wip[46].pnCode[4] := 0;
   hmiStns[4].wip[46].pnCode[5] := 0;
   hmiStns[4].wip[46].pnCode[6] := 0;
   hmiStns[4].wip[46].pnCode[7] := 0;
   hmiStns[4].wip[47].wipCode := -1;
   hmiStns[4].wip[47].pnCode[0] := 0;
   hmiStns[4].wip[47].pnCode[1] := 0;
   hmiStns[4].wip[47].pnCode[2] := 0;
   hmiStns[4].wip[47].pnCode[3] := 0;
   hmiStns[4].wip[47].pnCode[4] := 0;
   hmiStns[4].wip[47].pnCode[5] := 0;
   hmiStns[4].wip[47].pnCode[6] := 0;
   hmiStns[4].wip[47].pnCode[7] := 0;
   hmiStns[4].wip[48].wipCode := -1;
   hmiStns[4].wip[48].pnCode[0] := 0;
   hmiStns[4].wip[48].pnCode[1] := 0;
   hmiStns[4].wip[48].pnCode[2] := 0;
   hmiStns[4].wip[48].pnCode[3] := 0;
   hmiStns[4].wip[48].pnCode[4] := 0;
   hmiStns[4].wip[48].pnCode[5] := 0;
   hmiStns[4].wip[48].pnCode[6] := 0;
   hmiStns[4].wip[48].pnCode[7] := 0;
   hmiStns[4].wip[49].wipCode := -1;
   hmiStns[4].wip[49].pnCode[0] := 0;
   hmiStns[4].wip[49].pnCode[1] := 0;
   hmiStns[4].wip[49].pnCode[2] := 0;
   hmiStns[4].wip[49].pnCode[3] := 0;
   hmiStns[4].wip[49].pnCode[4] := 0;
   hmiStns[4].wip[49].pnCode[5] := 0;
   hmiStns[4].wip[49].pnCode[6] := 0;
   hmiStns[4].wip[49].pnCode[7] := 0;
END_DATA_BLOCK

// folder: Global Data

DATA_BLOCK "HMI Data: Warehouse HMI"   // DB2
{ S7_Optimized_Access := 'TRUE' }
VERSION : 0.1
   VAR
      barcode : "Barcode Screen";
      networkHealth : "Network Health Screen";
      partCall : "Part Call Screen";
      screenNumber : Int := 1;
      settings : "Settings";
      simStations : "Simulated Stations";
      tableNav : "Nav Bar Data: PLC";
      pop_up : "Pop Ups";
      settings_meta : "Setting Meta Data";
   END_VAR
BEGIN
END_DATA_BLOCK

